// Mitsubishi GX Works2 project: KotelnyaPLC   PLC: FX3U/FX3UC (continued)
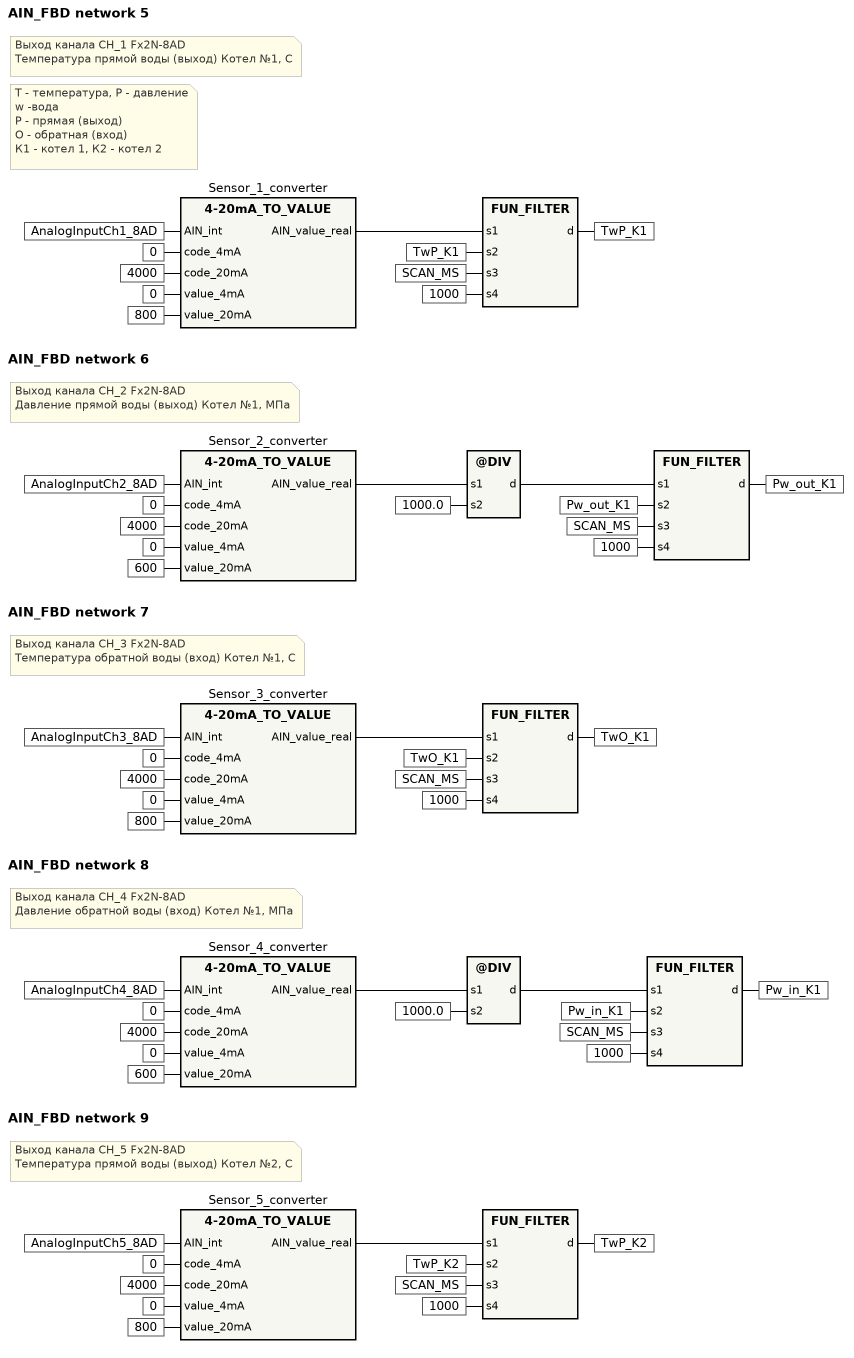
(* [picture p14: structured ladder/FBD of AIN_FBD, networks 5 to 9] *)
(* network 5 *)
(* Выход канала CH_1 Fx2N-8AD / Температура прямой воды (выход) Котел №1, С *)
(* T - температура, P - давление / w -вода / P - прямая (выход) / O - обратная (вход) / К1 - котел 1, К2 - котел 2 *)
Sensor_1_converter(AIN_int := AnalogInputCh1_8AD, code_4mA := 0, code_20mA := 4000, value_4mA := 0, value_20mA := 800);
TwP_K1 := FUN_FILTER(Sensor_1_converter.AIN_value_real, TwP_K1, SCAN_MS, 1000);
(* network 6 *)
(* Выход канала CH_2 Fx2N-8AD / Давление прямой воды (выход) Котел №1, МПа *)
Sensor_2_converter(AIN_int := AnalogInputCh2_8AD, code_4mA := 0, code_20mA := 4000, value_4mA := 0, value_20mA := 600);
Pw_out_K1 := FUN_FILTER(@DIV(Sensor_2_converter.AIN_value_real, 1000.0), Pw_out_K1, SCAN_MS, 1000);
(* network 7 *)
(* Выход канала CH_3 Fx2N-8AD / Температура обратной воды (вход) Котел №1, C *)
Sensor_3_converter(AIN_int := AnalogInputCh3_8AD, code_4mA := 0, code_20mA := 4000, value_4mA := 0, value_20mA := 800);
TwO_K1 := FUN_FILTER(Sensor_3_converter.AIN_value_real, TwO_K1, SCAN_MS, 1000);
(* network 8 *)
(* Выход канала CH_4 Fx2N-8AD / Давление обратной воды (вход) Котел №1, МПа *)
Sensor_4_converter(AIN_int := AnalogInputCh4_8AD, code_4mA := 0, code_20mA := 4000, value_4mA := 0, value_20mA := 600);
Pw_in_K1 := FUN_FILTER(@DIV(Sensor_4_converter.AIN_value_real, 1000.0), Pw_in_K1, SCAN_MS, 1000);
(* network 9 *)
(* Выход канала CH_5 Fx2N-8AD / Температура прямой воды (выход) Котел №2, С *)
Sensor_5_converter(AIN_int := AnalogInputCh5_8AD, code_4mA := 0, code_20mA := 4000, value_4mA := 0, value_20mA := 800);
TwP_K2 := FUN_FILTER(Sensor_5_converter.AIN_value_real, TwP_K2, SCAN_MS, 1000);
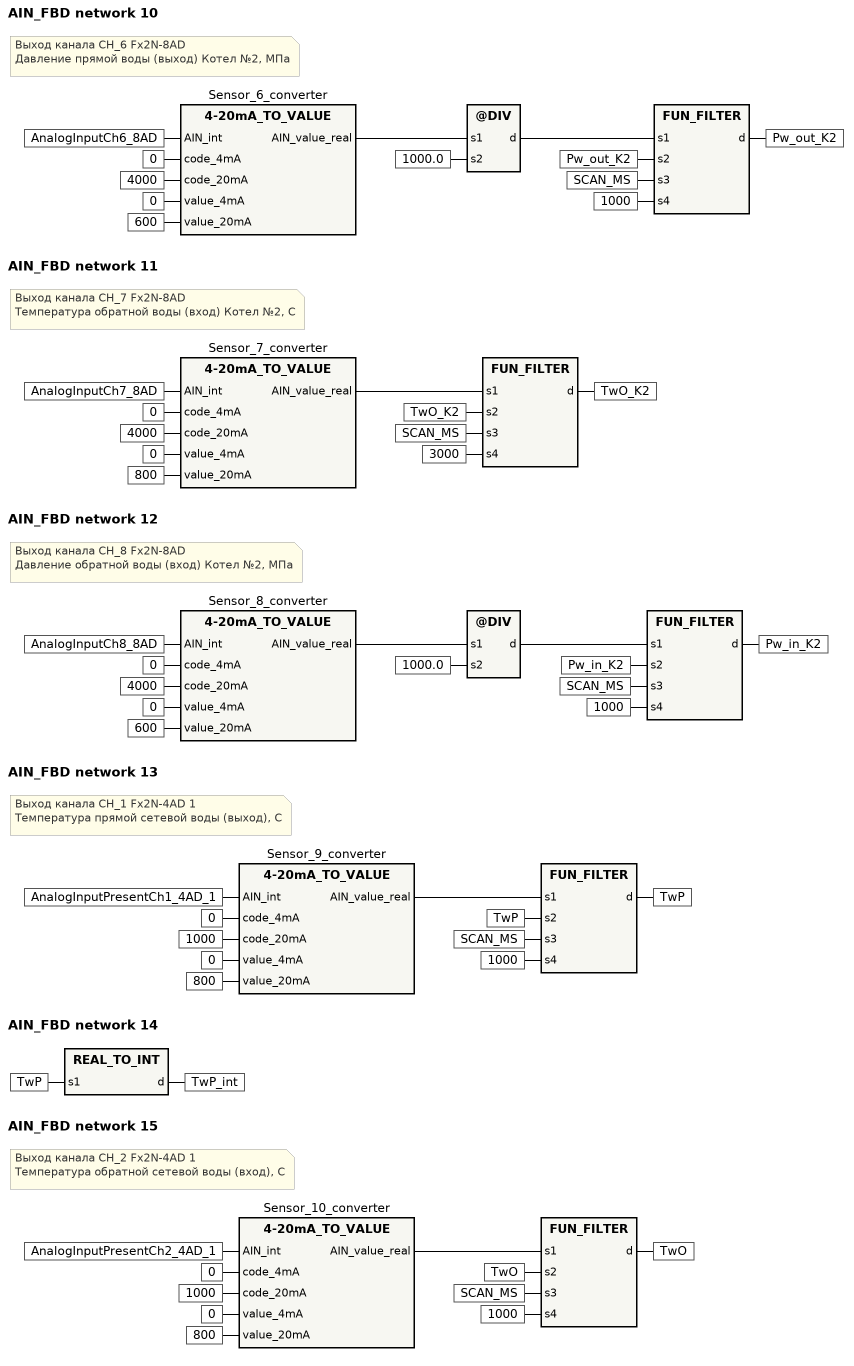
(* network 10 *)
(* Выход канала CH_6 Fx2N-8AD / Давление прямой воды (выход) Котел №2, МПа *)
Sensor_6_converter(AIN_int := AnalogInputCh6_8AD, code_4mA := 0, code_20mA := 4000, value_4mA := 0, value_20mA := 600);
Pw_out_K2 := FUN_FILTER(@DIV(Sensor_6_converter.AIN_value_real, 1000.0), Pw_out_K2, SCAN_MS, 1000);
(* network 11 *)
(* Выход канала CH_7 Fx2N-8AD / Температура обратной воды (вход) Котел №2, C *)
Sensor_7_converter(AIN_int := AnalogInputCh7_8AD, code_4mA := 0, code_20mA := 4000, value_4mA := 0, value_20mA := 800);
TwO_K2 := FUN_FILTER(Sensor_7_converter.AIN_value_real, TwO_K2, SCAN_MS, 3000);
(* network 12 *)
(* Выход канала CH_8 Fx2N-8AD / Давление обратной воды (вход) Котел №2, МПа *)
Sensor_8_converter(AIN_int := AnalogInputCh8_8AD, code_4mA := 0, code_20mA := 4000, value_4mA := 0, value_20mA := 600);
Pw_in_K2 := FUN_FILTER(@DIV(Sensor_8_converter.AIN_value_real, 1000.0), Pw_in_K2, SCAN_MS, 1000);
(* network 13 *)
(* Выход канала CH_1 Fx2N-4AD 1 / Температура прямой сетевой воды (выход), C *)
Sensor_9_converter(AIN_int := AnalogInputPresentCh1_4AD_1, code_4mA := 0, code_20mA := 1000, value_4mA := 0, value_20mA := 800);
TwP := FUN_FILTER(Sensor_9_converter.AIN_value_real, TwP, SCAN_MS, 1000);
(* network 14 *)
TwP_int := REAL_TO_INT(TwP);
(* network 15 *)
(* Выход канала CH_2 Fx2N-4AD 1 / Температура обратной сетевой воды (вход), C *)
Sensor_10_converter(AIN_int := AnalogInputPresentCh2_4AD_1, code_4mA := 0, code_20mA := 1000, value_4mA := 0, value_20mA := 800);
TwO := FUN_FILTER(Sensor_10_converter.AIN_value_real, TwO, SCAN_MS, 1000);
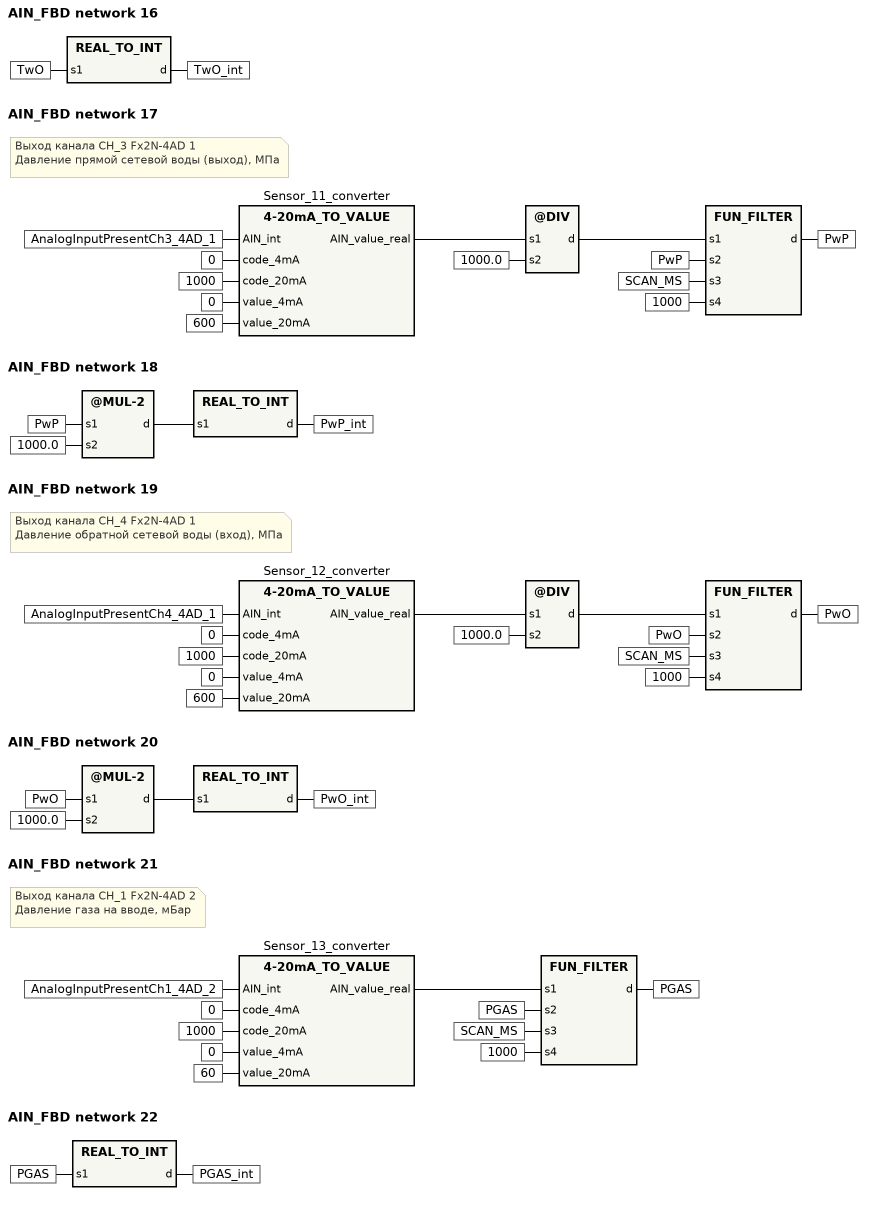
(* network 16 *)
TwO_int := REAL_TO_INT(TwO);
(* network 17 *)
(* Выход канала CH_3 Fx2N-4AD 1 / Давление прямой сетевой воды (выход), МПа *)
Sensor_11_converter(AIN_int := AnalogInputPresentCh3_4AD_1, code_4mA := 0, code_20mA := 1000, value_4mA := 0, value_20mA := 600);
PwP := FUN_FILTER(@DIV(Sensor_11_converter.AIN_value_real, 1000.0), PwP, SCAN_MS, 1000);
(* network 18 *)
PwP_int := REAL_TO_INT(@MUL-2(PwP, 1000.0));
(* network 19 *)
(* Выход канала CH_4 Fx2N-4AD 1 / Давление обратной сетевой воды (вход), МПа *)
Sensor_12_converter(AIN_int := AnalogInputPresentCh4_4AD_1, code_4mA := 0, code_20mA := 1000, value_4mA := 0, value_20mA := 600);
PwO := FUN_FILTER(@DIV(Sensor_12_converter.AIN_value_real, 1000.0), PwO, SCAN_MS, 1000);
(* network 20 *)
PwO_int := REAL_TO_INT(@MUL-2(PwO, 1000.0));
(* network 21 *)
(* Выход канала CH_1 Fx2N-4AD 2 / Давление газа на вводе, мБар *)
Sensor_13_converter(AIN_int := AnalogInputPresentCh1_4AD_2, code_4mA := 0, code_20mA := 1000, value_4mA := 0, value_20mA := 60);
PGAS := FUN_FILTER(Sensor_13_converter.AIN_value_real, PGAS, SCAN_MS, 1000);
(* network 22 *)
PGAS_int := REAL_TO_INT(PGAS);
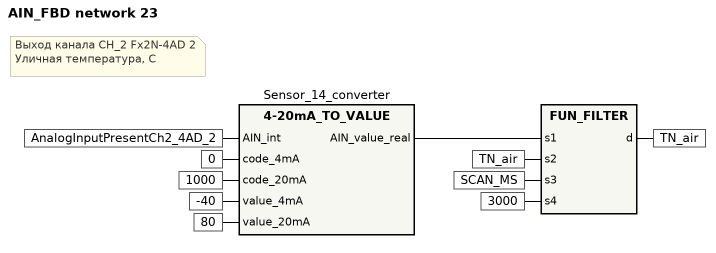
(* network 23 *)
(* Выход канала CH_2 Fx2N-4AD 2 / Уличная температура, С *)
Sensor_14_converter(AIN_int := AnalogInputPresentCh2_4AD_2, code_4mA := 0, code_20mA := 1000, value_4mA := -40, value_20mA := 80);
TN_air := FUN_FILTER(Sensor_14_converter.AIN_value_real, TN_air, SCAN_MS, 3000);
END_PROGRAM

FUNCTION_BLOCK 4-20mA_TO_VALUE
VAR_INPUT
  AIN_int : INT;
  code_4mA : INT;
  code_20mA : INT;
  value_4mA : INT;
  value_20mA : INT;
END_VAR
VAR
  code_4mA_real : REAL;
  code_20mA_real : REAL;
  value_4mA_real : REAL;
  value_20mA_real : REAL;
  AIN_real : REAL;
END_VAR
VAR_OUTPUT
  AIN_value_real : REAL;
END_VAR
VAR
  k1_real : REAL;
  c1_real : REAL;
END_VAR
(* structured ladder/FBD written out as ST: instructions are called as NAME(EN, inputs, outputs); _pN, _eN, _tN stand for wires *)
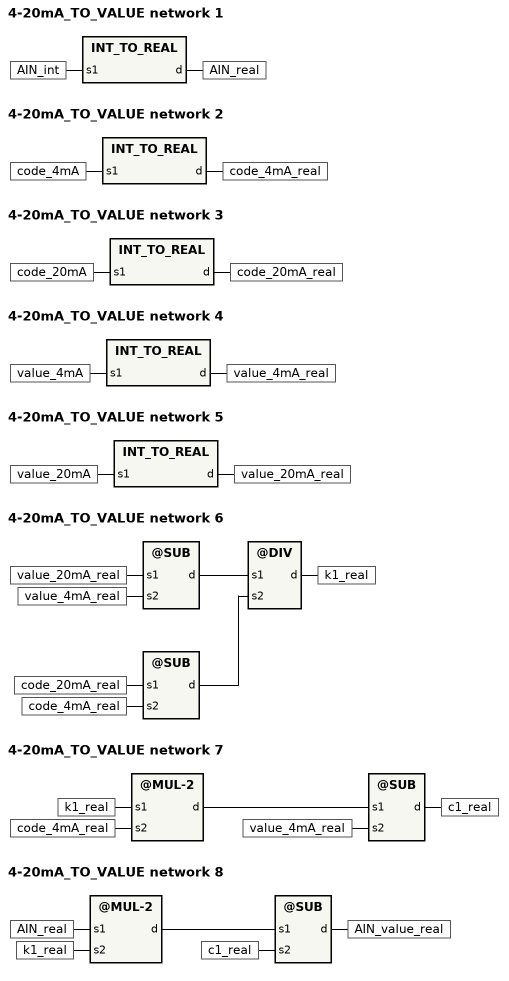
(* network 1 *)
AIN_real := INT_TO_REAL(AIN_int);
(* network 2 *)
code_4mA_real := INT_TO_REAL(code_4mA);
(* network 3 *)
code_20mA_real := INT_TO_REAL(code_20mA);
(* network 4 *)
value_4mA_real := INT_TO_REAL(value_4mA);
(* network 5 *)
value_20mA_real := INT_TO_REAL(value_20mA);
(* network 6 *)
k1_real := @DIV(@SUB(value_20mA_real, value_4mA_real), @SUB(code_20mA_real, code_4mA_real));
(* network 7 *)
c1_real := @SUB(@MUL-2(k1_real, code_4mA_real), value_4mA_real);
(* network 8 *)
AIN_value_real := @SUB(@MUL-2(AIN_real, k1_real), c1_real);
END_FUNCTION_BLOCK

FUNCTION_BLOCK KOTEL
VAR_INPUT
  Active_main : BOOL;  (* Активировать котел как главный *)
END_VAR
VAR_OUTPUT
  Alarm : BOOL;  (* Авария котла *)
  Burner_2 : BOOL;  (* Большое горение *)
  Dop_kotel : BOOL;  (* Второй котел *)
END_VAR
VAR_INPUT
  P_Water_IN : REAL;  (* Давление воды на входе в котел *)
  P_Water_OUT : REAL;  (* Давление воды на выходе из котла *)
  P_Water_MAX : REAL;  (* Давление воды максимальное (на выходе) *)
  P_Water_MIN : REAL;  (* Давление воды минимальное (на входе) *)
  Alarm_GOR : BOOL;  (* Авария с горелки котла *)
END_VAR
VAR_OUTPUT
  Burner_1 : BOOL;  (* Малое горение *)
END_VAR
VAR_INPUT
  TS_Water_95C : BOOL;  (* Термостат на выходе *)
  TS_Water_90C : BOOL;  (* Термостат на выходе *)
  Pdn40 : BOOL;  (* Датчик давления в топке ДН40 *)
  T_Water_80 : REAL;  (* Температура воды установленная большое горение *)
  T_Water_86 : REAL;  (* Температура воды установленная малое горение *)
  T_Water_OUT : REAL;  (* Датчик температуры на выходе котла *)
END_VAR
VAR_OUTPUT
  Recirc_Pump : BOOL;  (* Насос рециркуляции *)
END_VAR
VAR_INPUT
  T_Water_IN : REAL;  (* Температура воды на входе в котел *)
  T_Water_65 : REAL;  (* Температура воды установленная точка росы *)
END_VAR
VAR
  TON_1 : TON;
END_VAR
VAR_OUTPUT
  F_ALARM_P : BOOL;  (* Авария по давлению *)
END_VAR
VAR
  F_P_STOP : BOOL;  (* Стоп горелок по давлению *)
END_VAR
VAR_INPUT
  Rst_Alarm : BOOL;  (* Сброс аварии *)
END_VAR
VAR
  TOF_1 : TOF;
END_VAR
VAR_INPUT
  T_Water_90 : REAL;  (* Температура воды установленная выключение котла *)
END_VAR
VAR_OUTPUT
  Alarm_T_Water_90 : BOOL;  (* Авария котла при температуре на выходе более 90С *)
END_VAR
VAR
  Alarm_Pdn40 : BOOL;  (* Авария по датчику ДН-40 взрыв в топке *)
  TON_2 : TON;
  TOF_2 : TOF;
END_VAR
VAR_INPUT
  T_Water_IN_main : REAL;  (* Температура воды обратная общая *)
  T_Water_IN_main_ust : REAL;  (* Температура воды обратная общая установленная *)
  T_Water_hist : REAL;  (* Гистерезис температуры на включение горения *)
END_VAR
VAR
  TOF_3 : TOF;
  TON_3 : TON;
END_VAR
VAR_INPUT
  Active_dop : BOOL;  (* Активировать котел как дополнительный *)
END_VAR
VAR
  TON_4 : TON;
  TON_5 : TON;
  TOF_4 : TOF;
END_VAR
VAR_INPUT
  OP_Kotel_disable : BOOL;  (* Отключение работы котла *)
  OP_Dop_kotel : BOOL;  (* Включение дополнительного котла принудительно *)
END_VAR
VAR_OUTPUT
  OP_ALARM_P_sec : INT;
END_VAR
VAR_INPUT
  OP_Big_Fire : REAL;  (* Уставка включения большого горения и Дополнительного котла *)
END_VAR
VAR
  Active : BOOL;
  Active_1 : BOOL;
  Active_2 : BOOL;
END_VAR
VAR_OUTPUT
  P_Water_IN_status : INT;
  P_Water_OUT_status : INT;
  Time_Dop_kotel_on_min : INT;  (* Минут до включения доп котла *)
  Time_Dop_kotel_off_min : INT;  (* Минут до отключения доп котла *)
  Dop_kotel_on : BOOL;  (* Флаг таймера включения доп котла *)
  Dop_kotel_off : BOOL;  (* Флаг таймера включения доп котла *)
END_VAR
(* structured ladder/FBD written out as ST: instructions are called as NAME(EN, inputs, outputs); _pN, _eN, _tN stand for wires *)
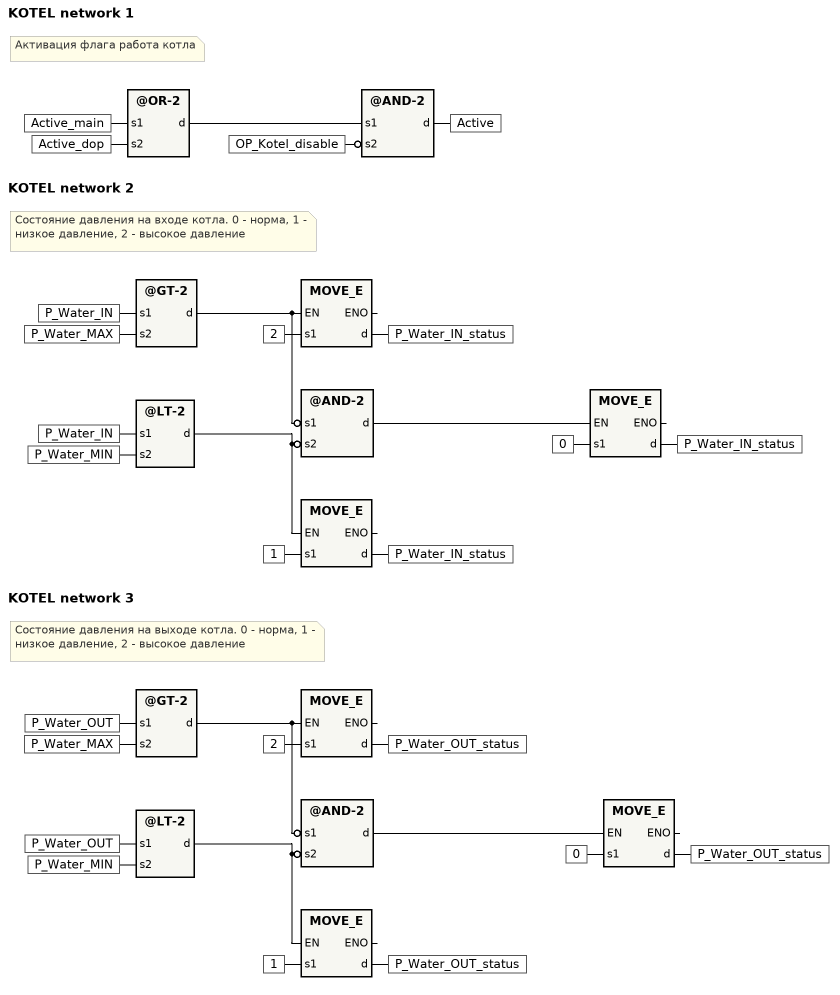
(* network 1 *)
(* Активация флага работа котла *)
Active := @AND-2(@OR-2(Active_main, Active_dop), NOT OP_Kotel_disable);
(* network 2 *)
(* Состояние давления на входе котла. 0 - норма, 1 - низкое давление, 2 - высокое давление *)
_p1 := @GT-2(P_Water_IN, P_Water_MAX);
MOVE_E(_p1, 2, P_Water_IN_status);
_p2 := @LT-2(P_Water_IN, P_Water_MIN);
MOVE_E(@AND-2(NOT _p1, NOT _p2), 0, P_Water_IN_status);
MOVE_E(_p2, 1, P_Water_IN_status);
(* network 3 *)
(* Состояние давления на выходе котла. 0 - норма, 1 - низкое давление, 2 - высокое давление *)
_p1 := @GT-2(P_Water_OUT, P_Water_MAX);
MOVE_E(_p1, 2, P_Water_OUT_status);
_p2 := @LT-2(P_Water_OUT, P_Water_MIN);
MOVE_E(@AND-2(NOT _p1, NOT _p2), 0, P_Water_OUT_status);
MOVE_E(_p2, 1, P_Water_OUT_status);
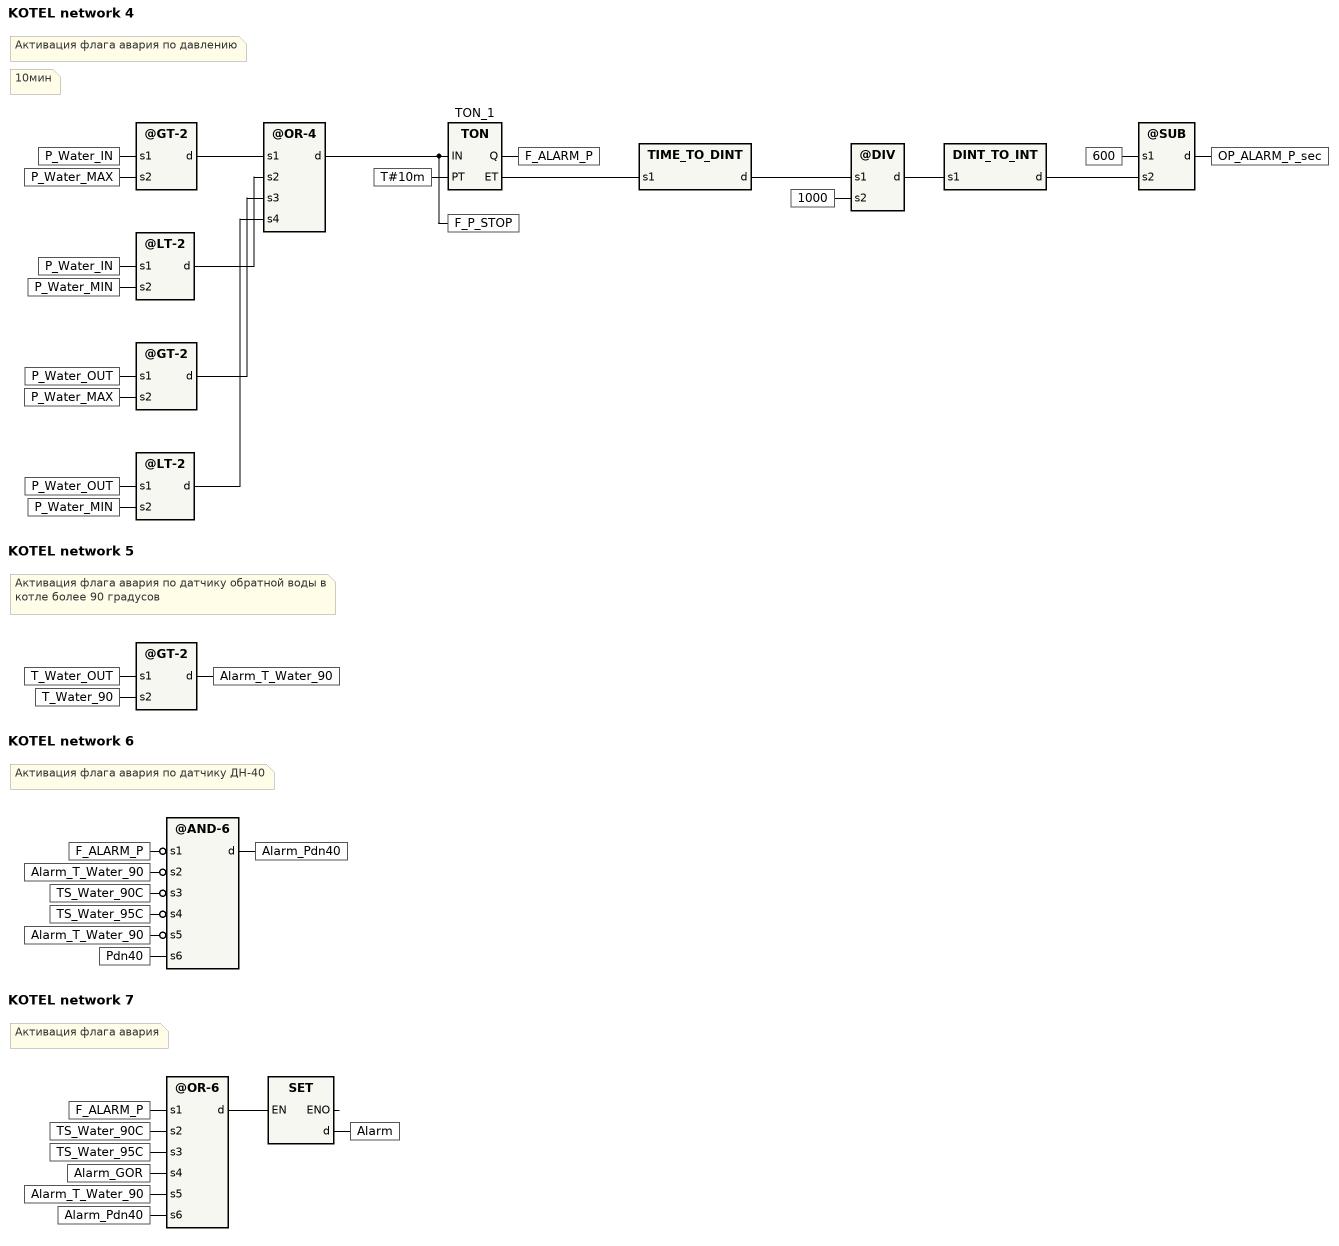
(* network 4 *)
(* Активация флага авария по давлению *)
(* 10мин *)
_p1 := @OR-4(@GT-2(P_Water_IN, P_Water_MAX), @LT-2(P_Water_IN, P_Water_MIN), @GT-2(P_Water_OUT, P_Water_MAX), @LT-2(P_Water_OUT, P_Water_MIN));
TON_1(IN := _p1, PT := T#10m, Q => F_ALARM_P);
OP_ALARM_P_sec := @SUB(600, DINT_TO_INT(@DIV(TIME_TO_DINT(TON_1.ET), 1000)));
F_P_STOP := _p1;
(* network 5 *)
(* Активация флага авария по датчику обратной воды в котле более 90 градусов *)
Alarm_T_Water_90 := @GT-2(T_Water_OUT, T_Water_90);
(* network 6 *)
(* Активация флага авария по датчику ДН-40 *)
Alarm_Pdn40 := @AND-6(NOT F_ALARM_P, NOT Alarm_T_Water_90, NOT TS_Water_90C, NOT TS_Water_95C, NOT Alarm_T_Water_90, Pdn40);
(* network 7 *)
(* Активация флага авария *)
SET(@OR-6(F_ALARM_P, TS_Water_90C, TS_Water_95C, Alarm_GOR, Alarm_T_Water_90, Alarm_Pdn40), Alarm);
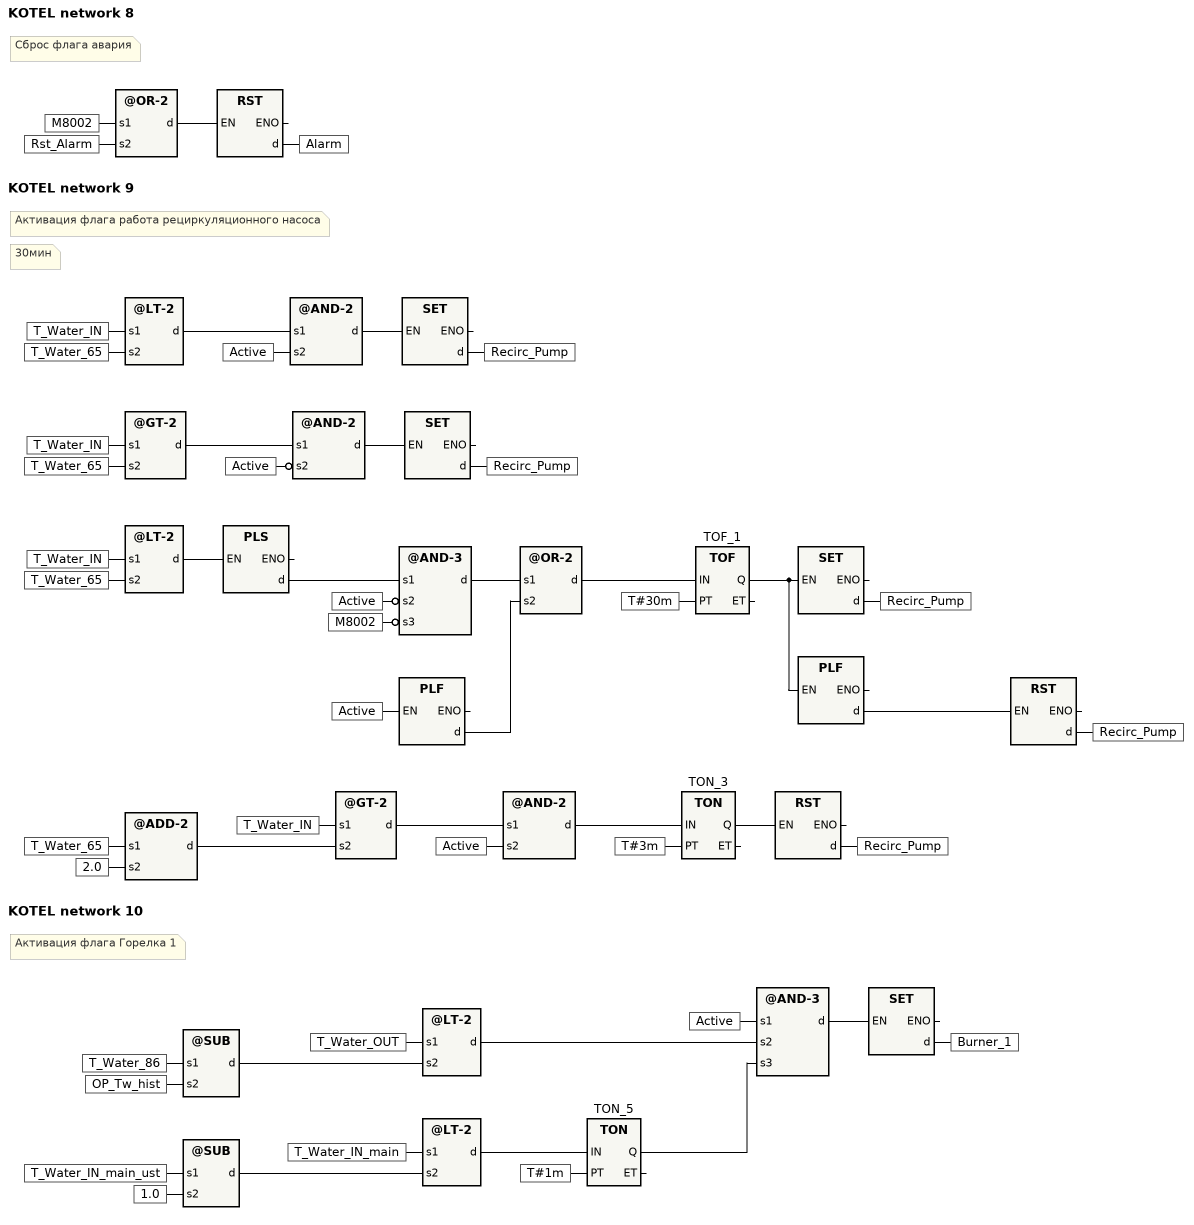
(* network 8 *)
(* Сброс флага авария *)
RST(@OR-2(M8002, Rst_Alarm), Alarm);
(* network 9 *)
(* Активация флага работа рециркуляционного насоса *)
(* 30мин *)
SET(@AND-2(@LT-2(T_Water_IN, T_Water_65), Active), Recirc_Pump);
SET(@AND-2(@GT-2(T_Water_IN, T_Water_65), NOT Active), Recirc_Pump);
PLS(@LT-2(T_Water_IN, T_Water_65), _t1);
PLF(Active, _t2);
TOF_1(IN := @OR-2(@AND-3(_t1, NOT Active, NOT M8002), _t2), PT := T#30m);
SET(TOF_1.Q, Recirc_Pump);
PLF(TOF_1.Q, _t3);
RST(_t3, Recirc_Pump);
TON_3(IN := @AND-2(@GT-2(T_Water_IN, @ADD-2(T_Water_65, 2.0)), Active), PT := T#3m);
RST(TON_3.Q, Recirc_Pump);
(* network 10 *)
(* Активация флага Горелка 1 *)
TON_5(IN := @LT-2(T_Water_IN_main, @SUB(T_Water_IN_main_ust, 1.0)), PT := T#1m);
SET(@AND-3(Active, @LT-2(T_Water_OUT, @SUB(T_Water_86, OP_Tw_hist)), TON_5.Q), Burner_1);
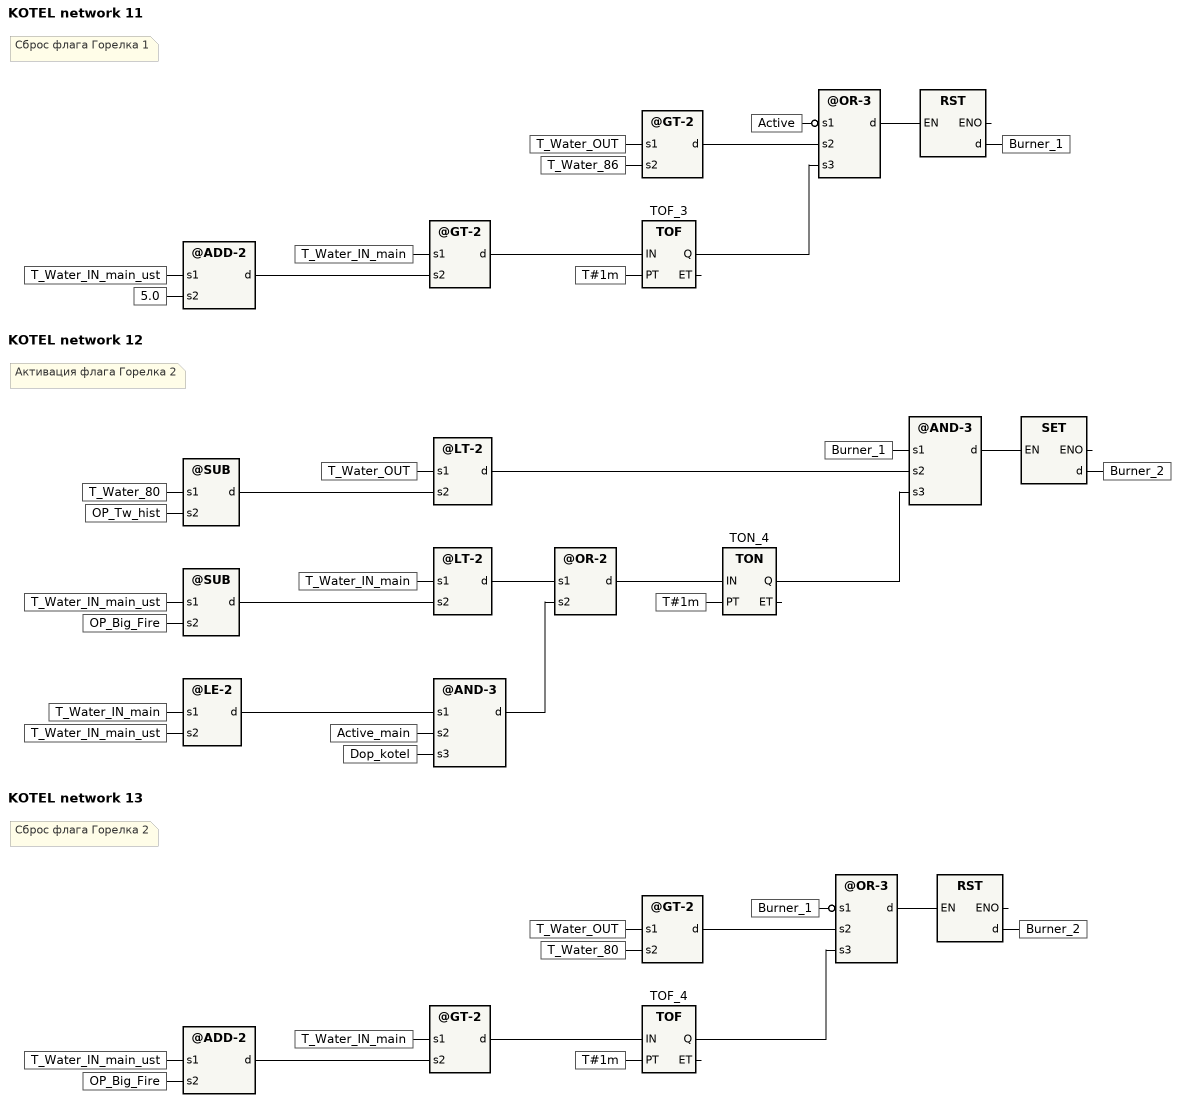
(* network 11 *)
(* Сброс флага Горелка 1 *)
TOF_3(IN := @GT-2(T_Water_IN_main, @ADD-2(T_Water_IN_main_ust, 5.0)), PT := T#1m);
RST(@OR-3(NOT Active, @GT-2(T_Water_OUT, T_Water_86), TOF_3.Q), Burner_1);
(* network 12 *)
(* Активация флага Горелка 2 *)
TON_4(IN := @OR-2(@LT-2(T_Water_IN_main, @SUB(T_Water_IN_main_ust, OP_Big_Fire)), @AND-3(@LE-2(T_Water_IN_main, T_Water_IN_main_ust), Active_main, Dop_kotel)), PT := T#1m);
SET(@AND-3(Burner_1, @LT-2(T_Water_OUT, @SUB(T_Water_80, OP_Tw_hist)), TON_4.Q), Burner_2);
(* network 13 *)
(* Сброс флага Горелка 2 *)
TOF_4(IN := @GT-2(T_Water_IN_main, @ADD-2(T_Water_IN_main_ust, OP_Big_Fire)), PT := T#1m);
RST(@OR-3(NOT Burner_1, @GT-2(T_Water_OUT, T_Water_80), TOF_4.Q), Burner_2);
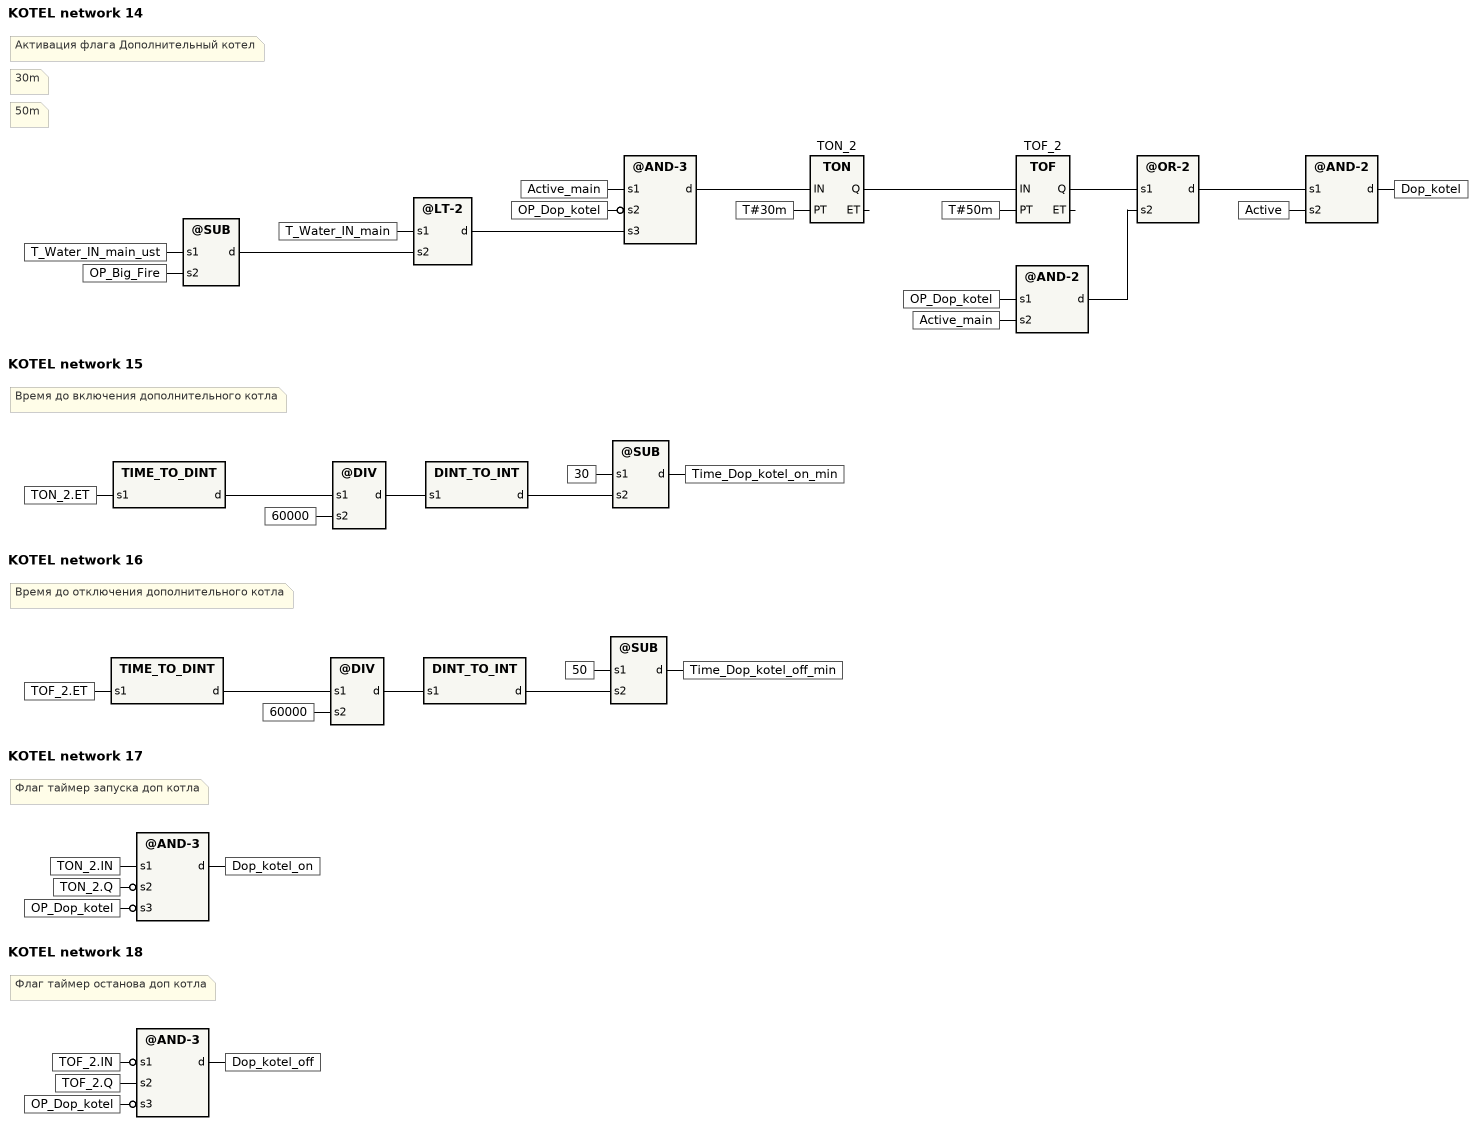
(* network 14 *)
(* Активация флага Дополнительный котел *)
(* 30m *)
(* 50m *)
TON_2(IN := @AND-3(Active_main, NOT OP_Dop_kotel, @LT-2(T_Water_IN_main, @SUB(T_Water_IN_main_ust, OP_Big_Fire))), PT := T#30m);
TOF_2(IN := TON_2.Q, PT := T#50m);
Dop_kotel := @AND-2(@OR-2(TOF_2.Q, @AND-2(OP_Dop_kotel, Active_main)), Active);
(* network 15 *)
(* Время до включения дополнительного котла *)
Time_Dop_kotel_on_min := @SUB(30, DINT_TO_INT(@DIV(TIME_TO_DINT(TON_2.ET), 60000)));
(* network 16 *)
(* Время до отключения дополнительного котла *)
Time_Dop_kotel_off_min := @SUB(50, DINT_TO_INT(@DIV(TIME_TO_DINT(TOF_2.ET), 60000)));
(* network 17 *)
(* Флаг таймер запуска доп котла *)
Dop_kotel_on := @AND-3(TON_2.IN, NOT TON_2.Q, NOT OP_Dop_kotel);
(* network 18 *)
(* Флаг таймер останова доп котла *)
Dop_kotel_off := @AND-3(NOT TOF_2.IN, TOF_2.Q, NOT OP_Dop_kotel);
END_FUNCTION_BLOCK

FUNCTION_BLOCK GRAPH
VAR_INPUT
  GRAPH_N : INT;  (* Номер графика *)
  DAY : INT;  (* Время суток День *)
  NIGHT : INT;  (* Время суток Ночь *)
  T_OUTDOOR : REAL;  (* Уличная температура *)
END_VAR
VAR_OUTPUT
  T_Water_IN_main_ust : REAL;  (* Температура обратной сетевой воды заданная *)
END_VAR
VAR
  F_NIGHT : BOOL;
  GRAPH_10 : REAL;  (* Температура обратной воды График 1 *)
  GRAPH_12 : REAL;  (* Температура обратной воды График 2 *)
  GRAPH_15 : REAL;  (* Температура обратной воды График 3 *)
  F_T_Water_IN_main_ust : REAL;
  Temp_Water_IN_main_ust : REAL;
END_VAR
VAR_INPUT
  T_CORR : INT;  (* Коррекция температуры обратной воды заданной *)
END_VAR
(* structured ladder/FBD written out as ST: instructions are called as NAME(EN, inputs, outputs); _pN, _eN, _tN stand for wires *)
